(* Logix 5000 project; controller PLC_MCC1300_75F1 vendor 1 type 14 code 166 rev 32.11; software revision 32.04; part 32 of 83 *)
(* tags used below, declared in another part *)
   BENCH_MASTERUP : ALIAS FOR I[73].6;
   I : INT[128];   // Local Input Updates Input Slot 2
   N14 : DINT[500];
   TD2_S_MOVIN : ALIAS FOR N14[256].5;
   TD2_S_MOVOUT : ALIAS FOR N14[257].5;
   TD3_N_MOVIN : ALIAS FOR N14[256].6;
   TD3_N_MOVOUT : ALIAS FOR N14[257].6;
   TD3_S_MOVIN : ALIAS FOR N14[256].7;
   TD3_S_MOVOUT : ALIAS FOR N14[257].7;
   TD4_N_MOVIN : ALIAS FOR N14[256].8;
   TD4_N_MOVOUT : ALIAS FOR N14[257].8;
   TD4_S_MOVIN : ALIAS FOR N14[256].9;
   TD4_S_MOVOUT : ALIAS FOR N14[257].9;
   TD5_N_MOVIN : ALIAS FOR N14[256].10;
   TD5_N_MOVOUT : ALIAS FOR N14[257].10;
   TD5_S_MOVIN : ALIAS FOR N14[256].11;
   TD5_S_MOVOUT : ALIAS FOR N14[257].11;
   TK3_N_MOVDN : ALIAS FOR N14[253].6;
   TK3_N_MOVIN : ALIAS FOR N14[254].6;
   TK3_N_MOVOUT : ALIAS FOR N14[255].6;
   TK3_N_MOVUP : ALIAS FOR N14[252].6;
   TK3_S_MOVDN : ALIAS FOR N14[253].7;
   TK3_S_MOVIN : ALIAS FOR N14[254].7;
   TK3_S_MOVOUT : ALIAS FOR N14[255].7;
   TK3_S_MOVUP : ALIAS FOR N14[252].7;
   TK4_N_MOVDN : ALIAS FOR N14[253].8;
   TK4_N_MOVIN : ALIAS FOR N14[254].8;
   TK4_N_MOVOUT : ALIAS FOR N14[255].8;
   TK4_N_MOVUP : ALIAS FOR N14[252].8;
   TK4_S_MOVDN : ALIAS FOR N14[253].9;
   TK4_S_MOVIN : ALIAS FOR N14[254].9;
   TK4_S_MOVOUT : ALIAS FOR N14[255].9;
   TK4_S_MOVUP : ALIAS FOR N14[252].9;
   TK5_N_MOVDN : ALIAS FOR N14[253].10;
   TK5_N_MOVIN : ALIAS FOR N14[254].10;
   TK5_N_MOVOUT : ALIAS FOR N14[255].10;
   TK5_N_MOVUP : ALIAS FOR N14[252].10;
   TK5_S_MOVDN : ALIAS FOR N14[253].11;
   TK5_S_MOVIN : ALIAS FOR N14[254].11;
   TK5_S_MOVOUT : ALIAS FOR N14[255].11;
   TK5_S_MOVUP : ALIAS FOR N14[252].11;
   TZ3_N_AUTO : ALIAS FOR N14[250].6;
   TZ3_N_MANL : ALIAS FOR N14[251].6;
   TZ3_S_AUTO : ALIAS FOR N14[250].7;
   TZ3_S_MANL : ALIAS FOR N14[251].7;
   TZ4_N_AUTO : ALIAS FOR N14[250].8;
   TZ4_N_MANL : ALIAS FOR N14[251].8;
   TZ4_S_AUTO : ALIAS FOR N14[250].9;
   TZ4_S_MANL : ALIAS FOR N14[251].9;
   TZ5_N_AUTO : ALIAS FOR N14[250].10;
   TZ5_N_MANL : ALIAS FOR N14[251].10;
   TZ5_S_AUTO : ALIAS FOR N14[250].11;
   TZ5_S_MANL : ALIAS FOR N14[251].11;
(* MainProgram, continued *)

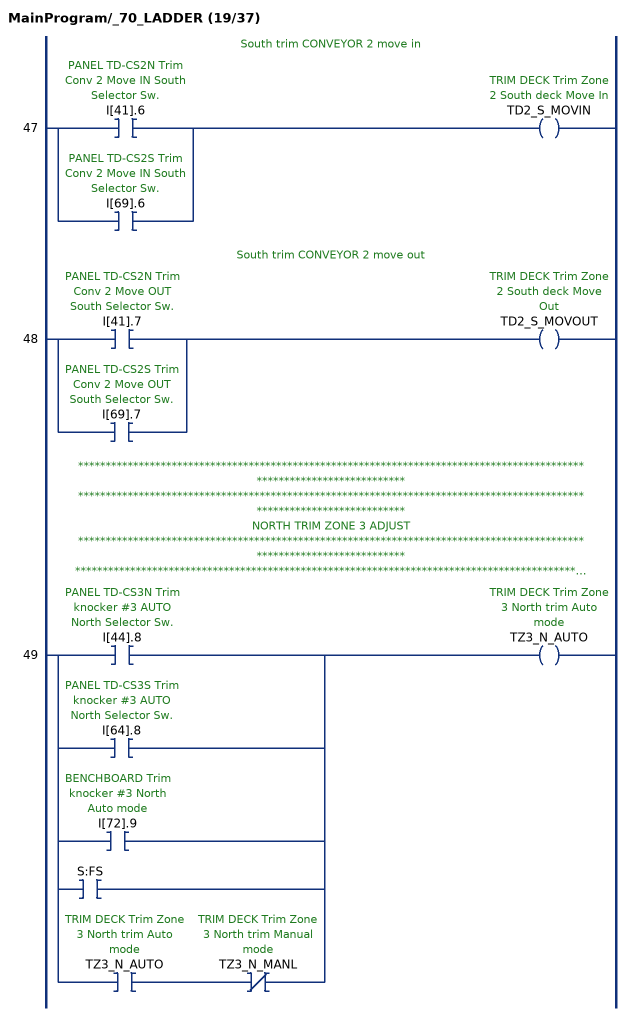
   [picture p450: MainProgram/_70_LADDER rungs 47-49]
   // South trim CONVEYOR 2 move in
   47: [XIC(I[41].6) ,XIC(I[69].6) ]OTE(TD2_S_MOVIN);
   // South trim CONVEYOR 2 move out
   48: [XIC(I[41].7) ,XIC(I[69].7) ]OTE(TD2_S_MOVOUT);
   // ***********************************************************************************************************************
   // ***********************************************************************************************************************
   //                                              NORTH TRIM ZONE 3 ADJUST
   // ***********************************************************************************************************************
   // ***********************************************************************************************************************
   // North trim knocker 3 auto mode
   49: [[XIC(I[44].8) ,XIC(I[64].8) ,XIC(I[72].9) ,XIC(S:FS) ] ,XIC(TZ3_N_AUTO) XIO(TZ3_N_MANL) ]OTE(TZ3_N_AUTO);
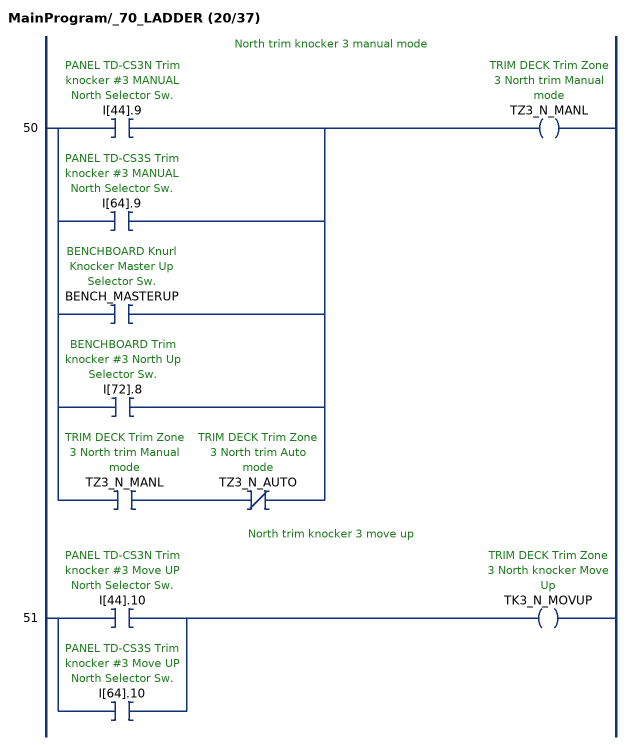
   // North trim knocker 3 manual mode
   50: [[XIC(I[44].9) ,XIC(I[64].9) ,XIC(BENCH_MASTERUP) ,XIC(I[72].8) ] ,XIC(TZ3_N_MANL) XIO(TZ3_N_AUTO) ]OTE(TZ3_N_MANL);
   // North trim knocker 3 move up
   51: [XIC(I[44].10) ,XIC(I[64].10) ]OTE(TK3_N_MOVUP);
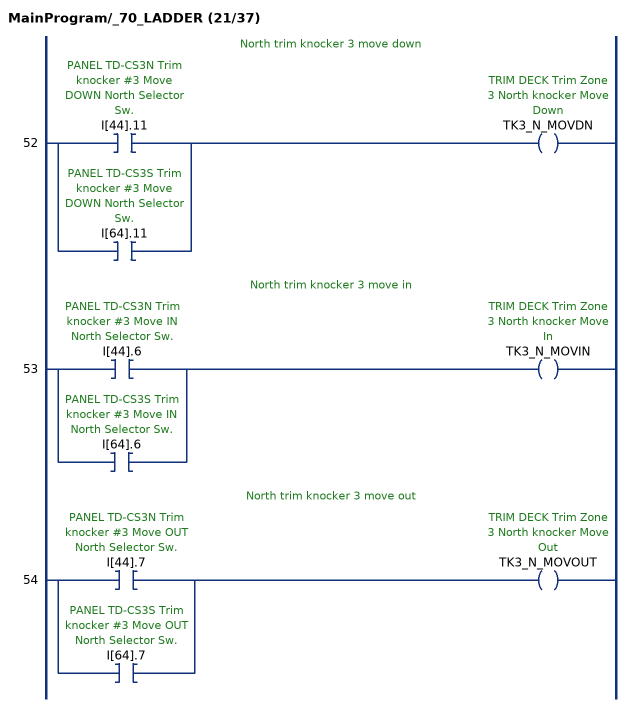
   // North trim knocker 3 move down
   52: [XIC(I[44].11) ,XIC(I[64].11) ]OTE(TK3_N_MOVDN);
   // North trim knocker 3 move in
   53: [XIC(I[44].6) ,XIC(I[64].6) ]OTE(TK3_N_MOVIN);
   // North trim knocker 3 move out
   54: [XIC(I[44].7) ,XIC(I[64].7) ]OTE(TK3_N_MOVOUT);
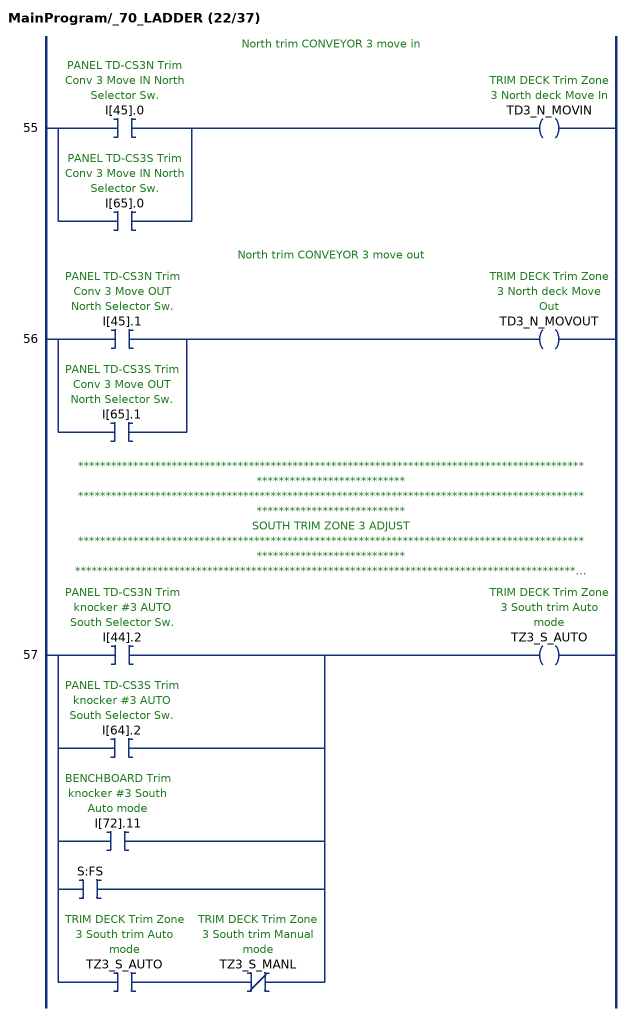
   // North trim CONVEYOR 3 move in
   55: [XIC(I[45].0) ,XIC(I[65].0) ]OTE(TD3_N_MOVIN);
   // North trim CONVEYOR 3 move out
   56: [XIC(I[45].1) ,XIC(I[65].1) ]OTE(TD3_N_MOVOUT);
   // ***********************************************************************************************************************
   // ***********************************************************************************************************************
   //                                              SOUTH TRIM ZONE 3 ADJUST
   // ***********************************************************************************************************************
   // ***********************************************************************************************************************
   // South trim knocker 3 auto mode
   57: [[XIC(I[44].2) ,XIC(I[64].2) ,XIC(I[72].11) ,XIC(S:FS) ] ,XIC(TZ3_S_AUTO) XIO(TZ3_S_MANL) ]OTE(TZ3_S_AUTO);
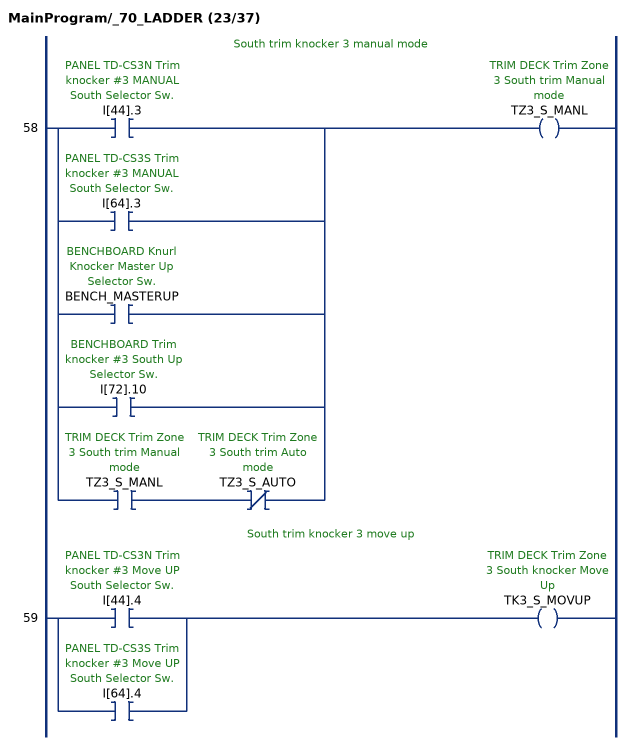
   // South trim knocker 3 manual mode
   58: [[XIC(I[44].3) ,XIC(I[64].3) ,XIC(BENCH_MASTERUP) ,XIC(I[72].10) ] ,XIC(TZ3_S_MANL) XIO(TZ3_S_AUTO) ]OTE(TZ3_S_MANL);
   // South trim knocker 3 move up
   59: [XIC(I[44].4) ,XIC(I[64].4) ]OTE(TK3_S_MOVUP);
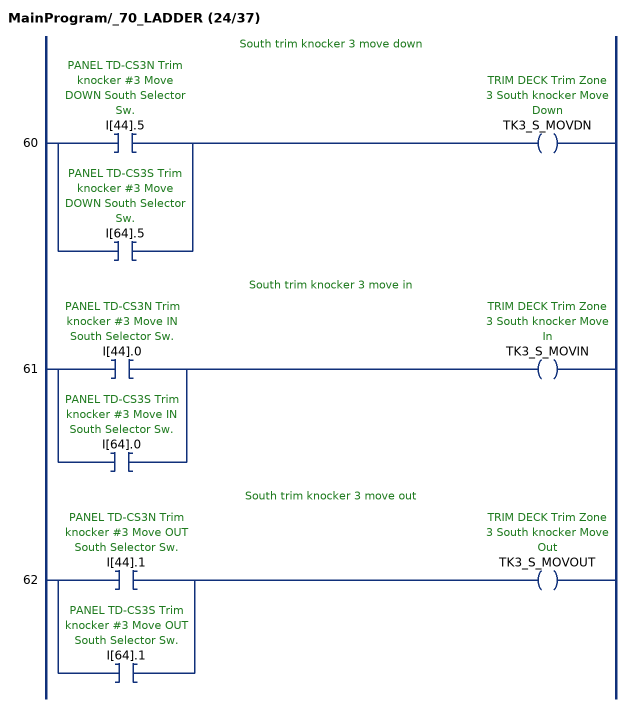
   // South trim knocker 3 move down
   60: [XIC(I[44].5) ,XIC(I[64].5) ]OTE(TK3_S_MOVDN);
   // South trim knocker 3 move in
   61: [XIC(I[44].0) ,XIC(I[64].0) ]OTE(TK3_S_MOVIN);
   // South trim knocker 3 move out
   62: [XIC(I[44].1) ,XIC(I[64].1) ]OTE(TK3_S_MOVOUT);
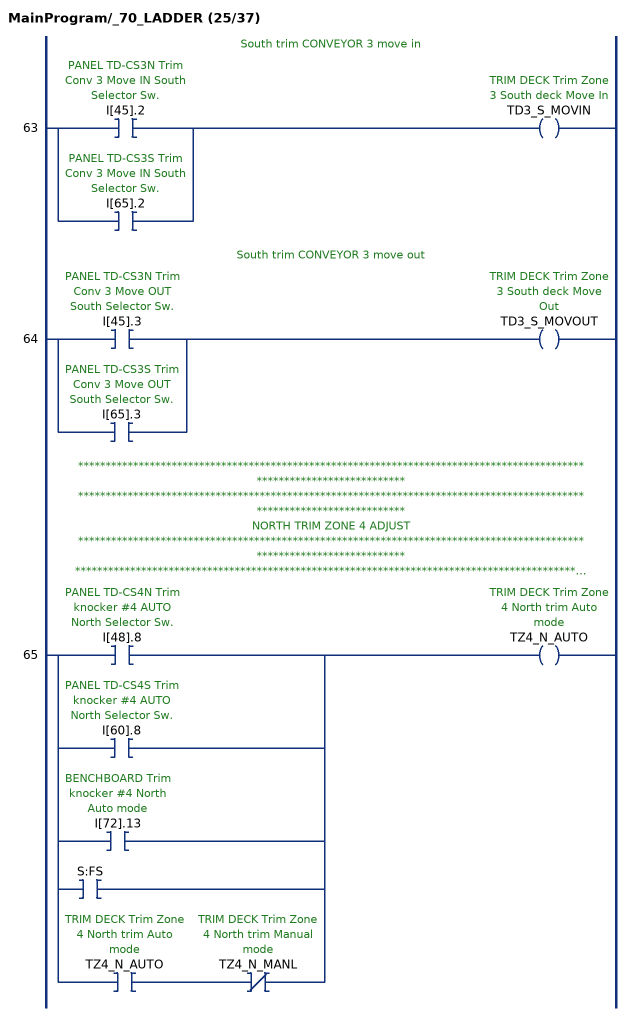
   // South trim CONVEYOR 3 move in
   63: [XIC(I[45].2) ,XIC(I[65].2) ]OTE(TD3_S_MOVIN);
   // South trim CONVEYOR 3 move out
   64: [XIC(I[45].3) ,XIC(I[65].3) ]OTE(TD3_S_MOVOUT);
   // ***********************************************************************************************************************
   // ***********************************************************************************************************************
   //                                              NORTH TRIM ZONE 4 ADJUST
   // ***********************************************************************************************************************
   // ***********************************************************************************************************************
   // North trim knocker 4 auto mode
   65: [[XIC(I[48].8) ,XIC(I[60].8) ,XIC(I[72].13) ,XIC(S:FS) ] ,XIC(TZ4_N_AUTO) XIO(TZ4_N_MANL) ]OTE(TZ4_N_AUTO);
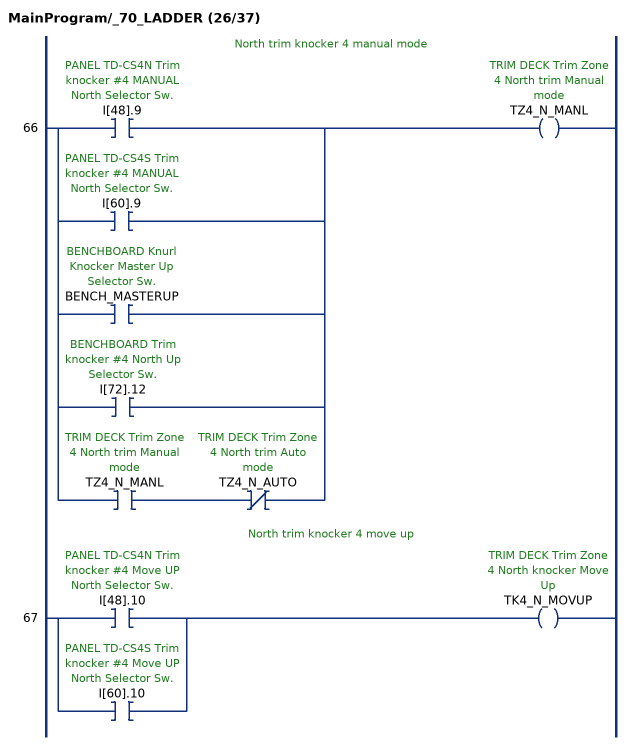
   // North trim knocker 4 manual mode
   66: [[XIC(I[48].9) ,XIC(I[60].9) ,XIC(BENCH_MASTERUP) ,XIC(I[72].12) ] ,XIC(TZ4_N_MANL) XIO(TZ4_N_AUTO) ]OTE(TZ4_N_MANL);
   // North trim knocker 4 move up
   67: [XIC(I[48].10) ,XIC(I[60].10) ]OTE(TK4_N_MOVUP);
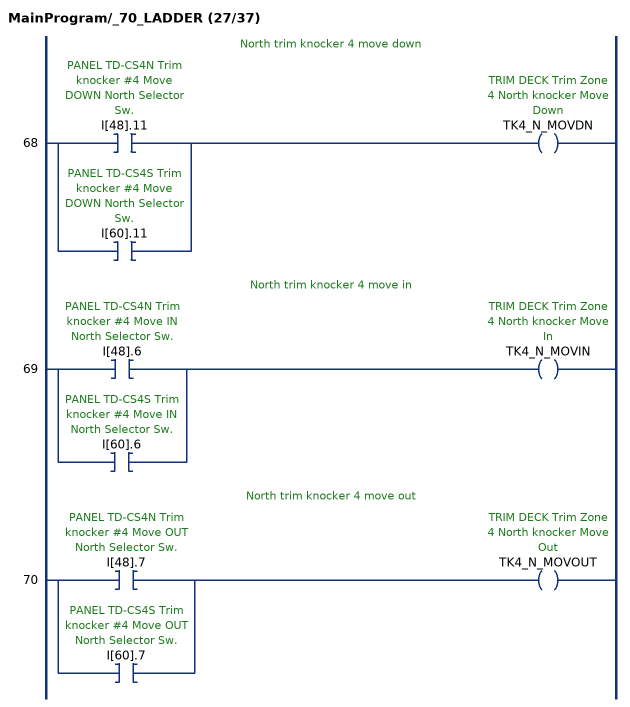
   // North trim knocker 4 move down
   68: [XIC(I[48].11) ,XIC(I[60].11) ]OTE(TK4_N_MOVDN);
   // North trim knocker 4 move in
   69: [XIC(I[48].6) ,XIC(I[60].6) ]OTE(TK4_N_MOVIN);
   // North trim knocker 4 move out
   70: [XIC(I[48].7) ,XIC(I[60].7) ]OTE(TK4_N_MOVOUT);
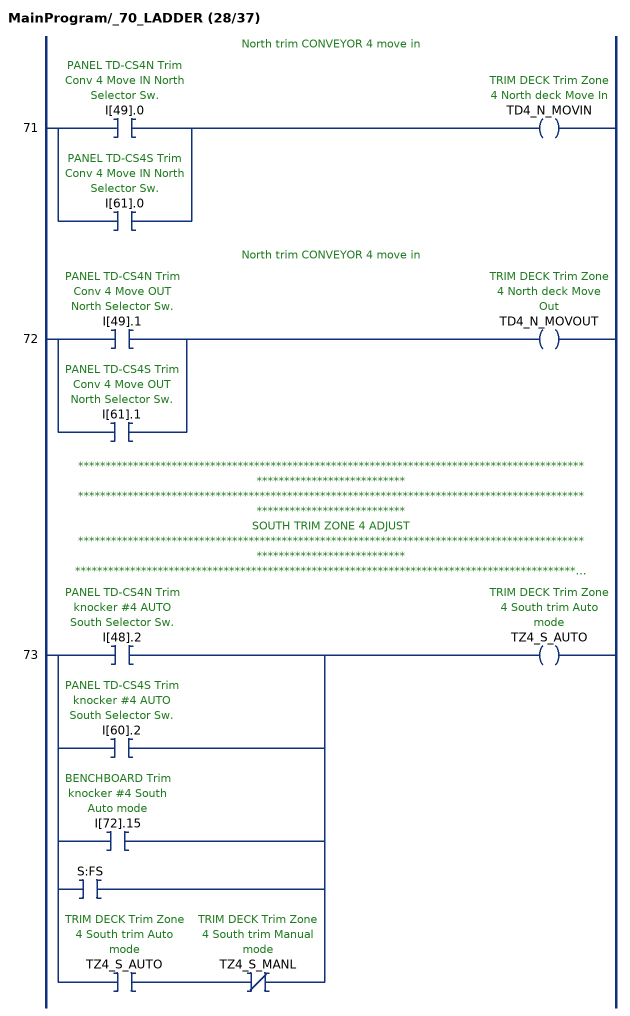
   // North trim CONVEYOR 4 move in
   71: [XIC(I[49].0) ,XIC(I[61].0) ]OTE(TD4_N_MOVIN);
   // North trim CONVEYOR 4 move in
   72: [XIC(I[49].1) ,XIC(I[61].1) ]OTE(TD4_N_MOVOUT);
   // ***********************************************************************************************************************
   // ***********************************************************************************************************************
   //                                              SOUTH TRIM ZONE 4 ADJUST
   // ***********************************************************************************************************************
   // ***********************************************************************************************************************
   // South trim knocker 4 auto mode
   73: [[XIC(I[48].2) ,XIC(I[60].2) ,XIC(I[72].15) ,XIC(S:FS) ] ,XIC(TZ4_S_AUTO) XIO(TZ4_S_MANL) ]OTE(TZ4_S_AUTO);
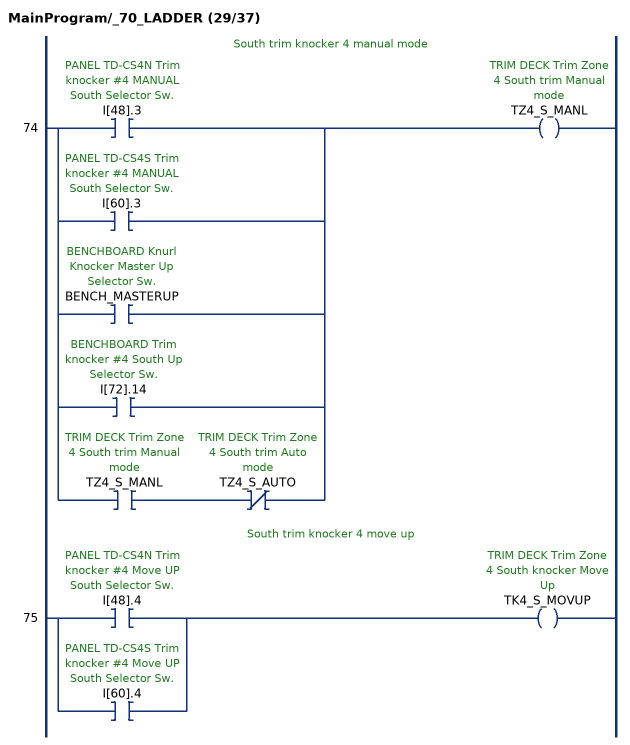
   // South trim knocker 4 manual mode
   74: [[XIC(I[48].3) ,XIC(I[60].3) ,XIC(BENCH_MASTERUP) ,XIC(I[72].14) ] ,XIC(TZ4_S_MANL) XIO(TZ4_S_AUTO) ]OTE(TZ4_S_MANL);
   // South trim knocker 4 move up
   75: [XIC(I[48].4) ,XIC(I[60].4) ]OTE(TK4_S_MOVUP);
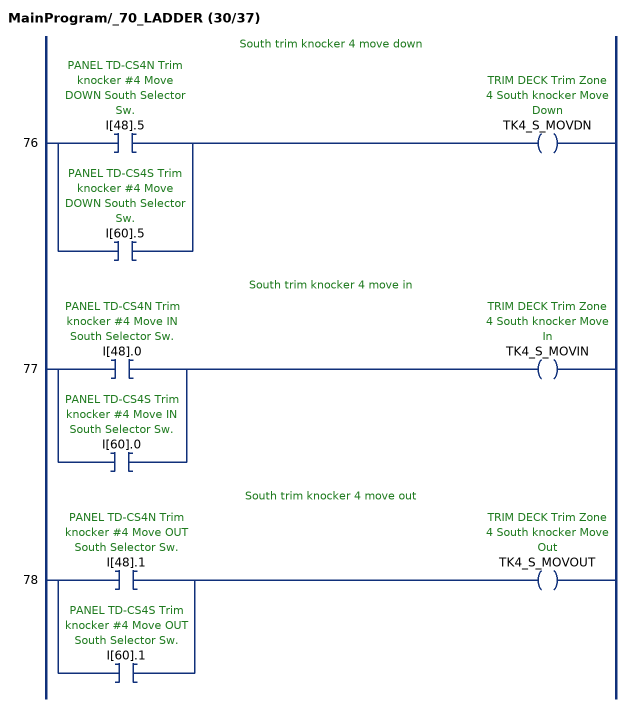
   // South trim knocker 4 move down
   76: [XIC(I[48].5) ,XIC(I[60].5) ]OTE(TK4_S_MOVDN);
   // South trim knocker 4 move in
   77: [XIC(I[48].0) ,XIC(I[60].0) ]OTE(TK4_S_MOVIN);
   // South trim knocker 4 move out
   78: [XIC(I[48].1) ,XIC(I[60].1) ]OTE(TK4_S_MOVOUT);
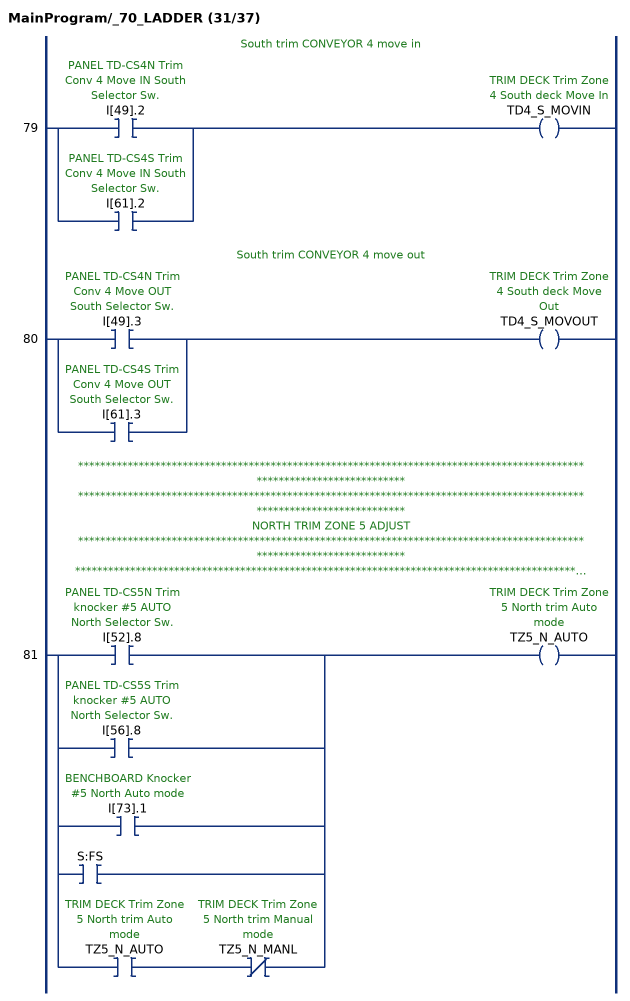
   // South trim CONVEYOR 4 move in
   79: [XIC(I[49].2) ,XIC(I[61].2) ]OTE(TD4_S_MOVIN);
   // South trim CONVEYOR 4 move out
   80: [XIC(I[49].3) ,XIC(I[61].3) ]OTE(TD4_S_MOVOUT);
   // ***********************************************************************************************************************
   // ***********************************************************************************************************************
   //                                              NORTH TRIM ZONE 5 ADJUST
   // ***********************************************************************************************************************
   // ***********************************************************************************************************************
   // North trim knocker 5 auto mode
   81: [[XIC(I[52].8) ,XIC(I[56].8) ,XIC(I[73].1) ,XIC(S:FS) ] ,XIC(TZ5_N_AUTO) XIO(TZ5_N_MANL) ]OTE(TZ5_N_AUTO);
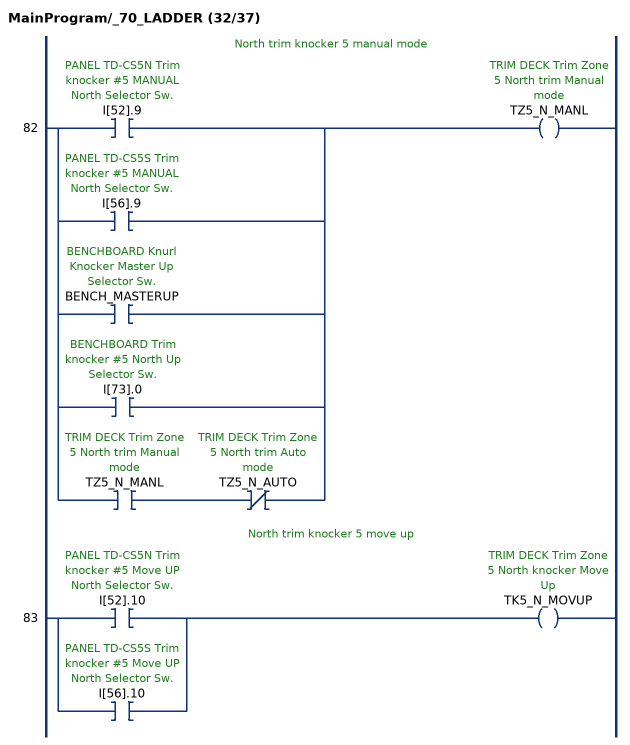
   // North trim knocker 5 manual mode
   82: [[XIC(I[52].9) ,XIC(I[56].9) ,XIC(BENCH_MASTERUP) ,XIC(I[73].0) ] ,XIC(TZ5_N_MANL) XIO(TZ5_N_AUTO) ]OTE(TZ5_N_MANL);
   // North trim knocker 5 move up
   83: [XIC(I[52].10) ,XIC(I[56].10) ]OTE(TK5_N_MOVUP);
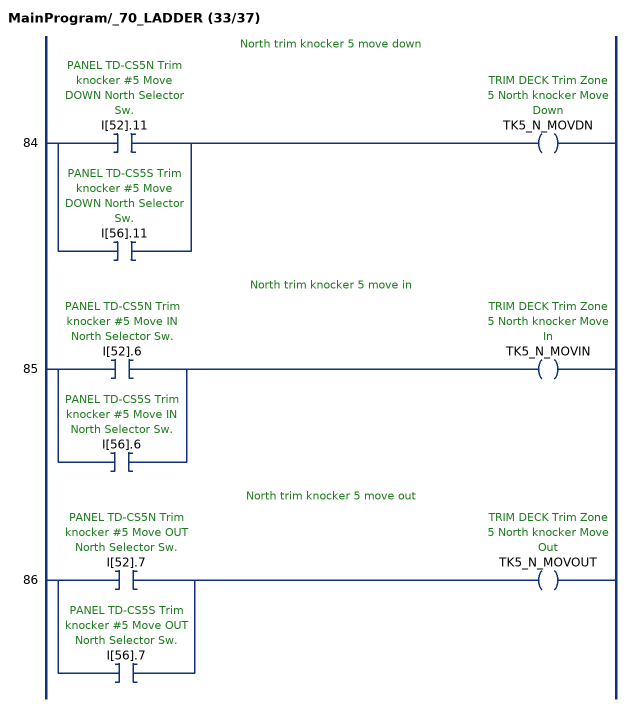
   // North trim knocker 5 move down
   84: [XIC(I[52].11) ,XIC(I[56].11) ]OTE(TK5_N_MOVDN);
   // North trim knocker 5 move in
   85: [XIC(I[52].6) ,XIC(I[56].6) ]OTE(TK5_N_MOVIN);
   // North trim knocker 5 move out
   86: [XIC(I[52].7) ,XIC(I[56].7) ]OTE(TK5_N_MOVOUT);
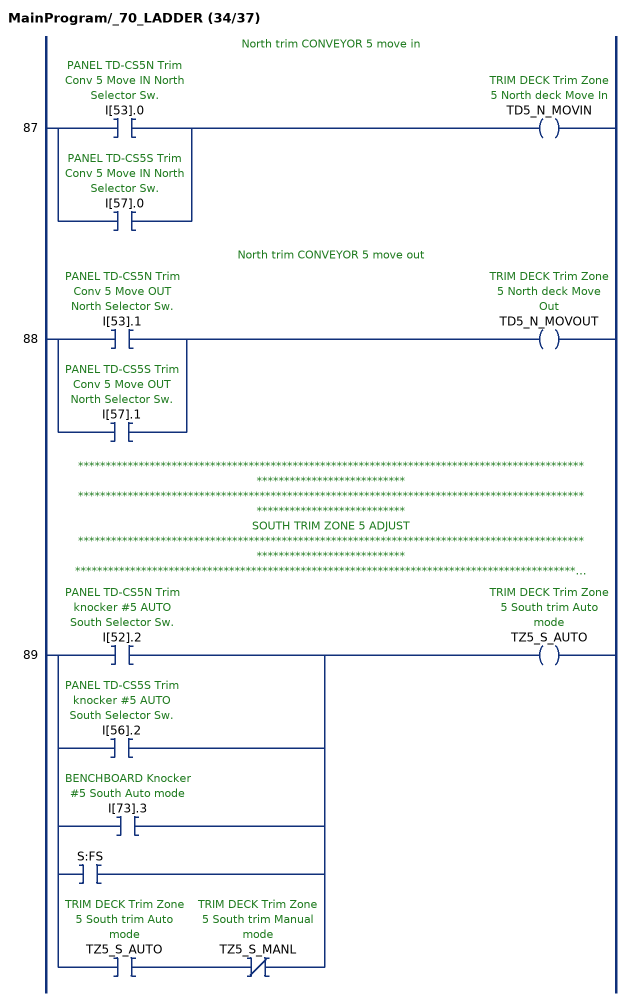
   // North trim CONVEYOR 5 move in
   87: [XIC(I[53].0) ,XIC(I[57].0) ]OTE(TD5_N_MOVIN);
   // North trim CONVEYOR 5 move out
   88: [XIC(I[53].1) ,XIC(I[57].1) ]OTE(TD5_N_MOVOUT);
   // ***********************************************************************************************************************
   // ***********************************************************************************************************************
   //                                              SOUTH TRIM ZONE 5 ADJUST
   // ***********************************************************************************************************************
   // ***********************************************************************************************************************
   // South trim knocker 5 auto mode
   89: [[XIC(I[52].2) ,XIC(I[56].2) ,XIC(I[73].3) ,XIC(S:FS) ] ,XIC(TZ5_S_AUTO) XIO(TZ5_S_MANL) ]OTE(TZ5_S_AUTO);
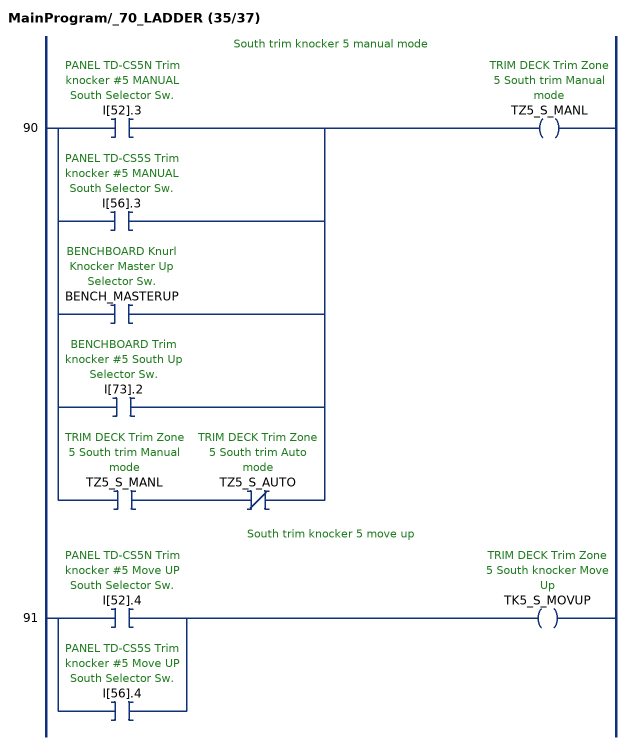
   // South trim knocker 5 manual mode
   90: [[XIC(I[52].3) ,XIC(I[56].3) ,XIC(BENCH_MASTERUP) ,XIC(I[73].2) ] ,XIC(TZ5_S_MANL) XIO(TZ5_S_AUTO) ]OTE(TZ5_S_MANL);
   // South trim knocker 5 move up
   91: [XIC(I[52].4) ,XIC(I[56].4) ]OTE(TK5_S_MOVUP);
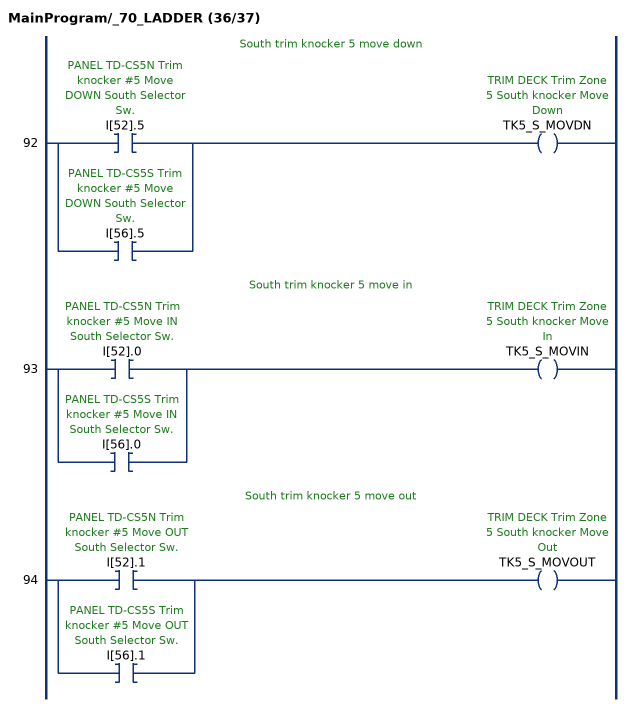
   // South trim knocker 5 move down
   92: [XIC(I[52].5) ,XIC(I[56].5) ]OTE(TK5_S_MOVDN);
   // South trim knocker 5 move in
   93: [XIC(I[52].0) ,XIC(I[56].0) ]OTE(TK5_S_MOVIN);
   // South trim knocker 5 move out
   94: [XIC(I[52].1) ,XIC(I[56].1) ]OTE(TK5_S_MOVOUT);
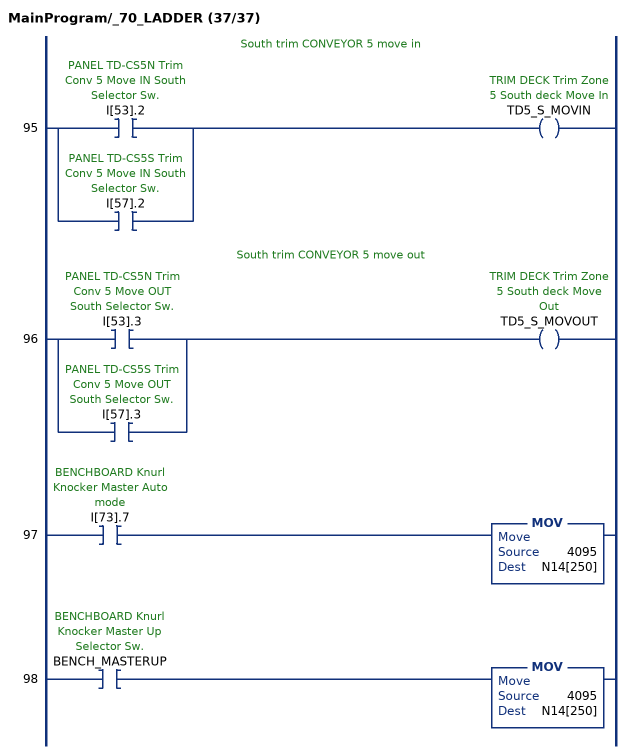
   // South trim CONVEYOR 5 move in
   95: [XIC(I[53].2) ,XIC(I[57].2) ]OTE(TD5_S_MOVIN);
   // South trim CONVEYOR 5 move out
   96: [XIC(I[53].3) ,XIC(I[57].3) ]OTE(TD5_S_MOVOUT);
   97: XIC(I[73].7)MOV(4095,N14[250]);
   98: XIC(BENCH_MASTERUP)MOV(4095,N14[250]);
END_ROUTINE
